// TIA Portal project "Pozycjoner_v7" (V15.1) (continued)
REGION Network 3: Line 1 is in or out range: 5mm around Y avg point
   #_w1 := #Enabled AND ((#Line1.Y1 < "DB_Average positions".Ranges.DiffX.Min) OR (#Line1.Y1 > "DB_Average positions".Ranges.DiffX.Max));
   IF #_w1 THEN #DiffResult := #Line1.Y1 - "DB_Average positions".AveragePosition.Y; END_IF;
   #SetCount1 := #_w1 AND NOT #Ptrig1;   // rising edge
   #Ptrig1 := #_w1;
   IF #Enabled AND ("DB_Average positions".Ranges.DiffX.Min <= #Line1.Y1) AND (#Line1.Y1 <= "DB_Average positions".Ranges.DiffX.Max) THEN
       #GeneralXavg := "DB_Drivers".X_AVG;
       #MoveToCenter_IR := TRUE;
   END_IF;
   IF #SetCount1 THEN
       #MainCounter := 1;
       #RECountLine3 := 0;
   END_IF;
END_REGION

REGION Network 4: Shift by difference value
   RUNG wire#powerrail
      { S7_Templates := "SrcType := Real" } GT_Contact(in1 := #DiffResult, in2 := 0.0)
      Sub(in1 := "DB_Average positions".AveragePosition.Y, in2 := #DiffResult, out => #ShiftDifValue)
   END_RUNG
   RUNG wire#powerrail
      { S7_Templates := "SrcType := Real" } LT_Contact(in1 := #DiffResult, in2 := 0.0)
      { S7_Templates := "SrcType := Real" } Abs(in := #DiffResult, out => #DiffResult)
      Add(in1 := "DB_Average positions".AveragePosition.Y, in2 := #DiffResult, out => #ShiftDifValue)
   END_RUNG
   // the same network as SCL:
   IF #DiffResult > 0.0 THEN
       #ShiftDifValue := "DB_Average positions".AveragePosition.Y - #DiffResult;
   END_IF;
   #_w1 := #DiffResult < 0.0;
   IF #_w1 THEN
       #DiffResult := ABS(#DiffResult);
       #ShiftDifValue := "DB_Average positions".AveragePosition.Y + #DiffResult;
   END_IF;
END_REGION

REGION Network 5: Movement to the new line: 3
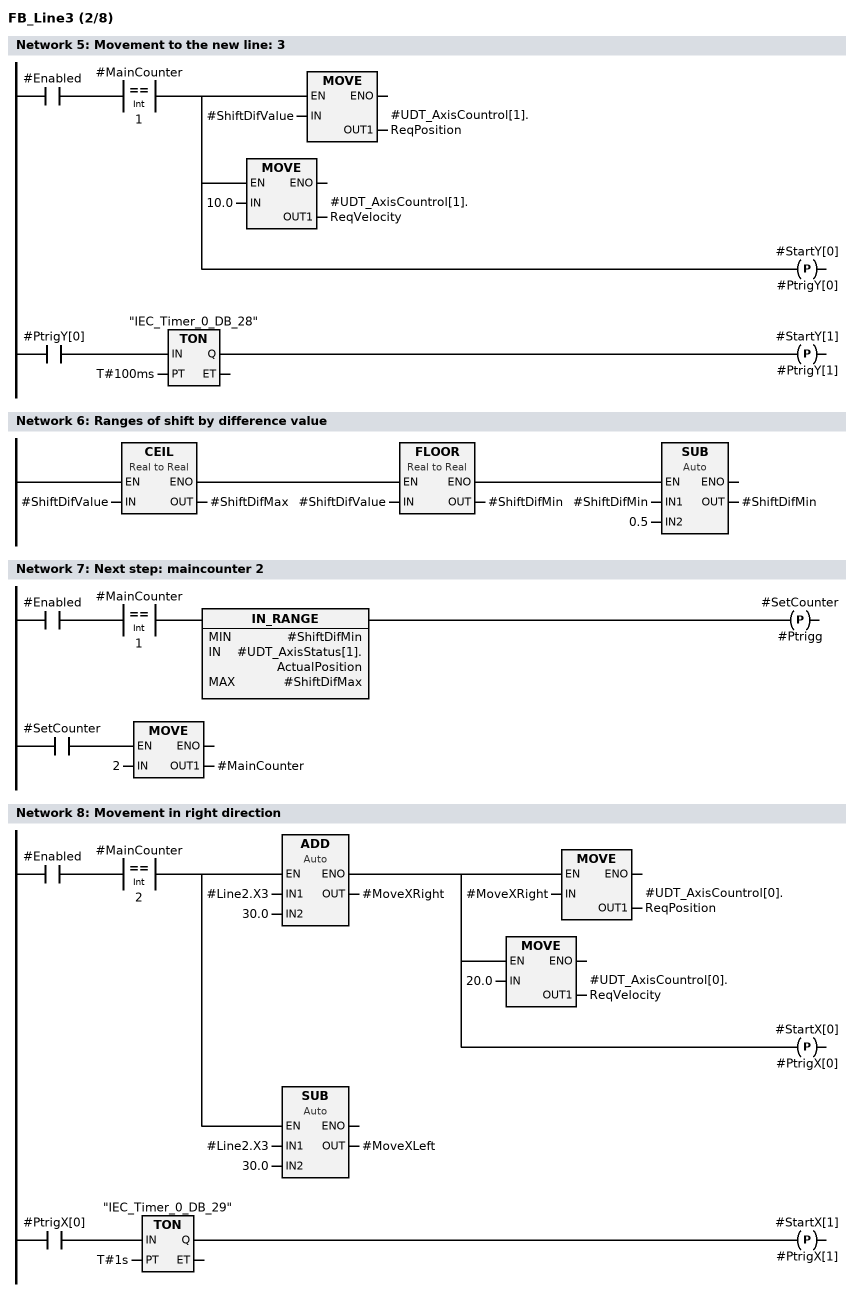
   #_w1 := #Enabled AND (#MainCounter = 1);
   IF #_w1 THEN
       #UDT_AxisCountrol[1].ReqPosition := #ShiftDifValue;
       #UDT_AxisCountrol[1].ReqVelocity := 10.0;
   END_IF;
   #StartY[0] := #_w1 AND NOT #PtrigY[0];   // rising edge
   #PtrigY[0] := #_w1;
   "IEC_Timer_0_DB_28".TON(IN := #PtrigY[0], PT := T#100ms);
   #StartY[1] := "IEC_Timer_0_DB_28".Q AND NOT #PtrigY[1];   // rising edge
   #PtrigY[1] := "IEC_Timer_0_DB_28".Q;
END_REGION

REGION Network 6: Ranges of shift by difference value
   #ShiftDifMax := CEIL(#ShiftDifValue);
   #ShiftDifMin := FLOOR(#ShiftDifValue);
   #ShiftDifMin := #ShiftDifMin - 0.5;
END_REGION

REGION Network 7: Next step: maincounter 2
   #_w1 := #Enabled AND (#MainCounter = 1) AND (#ShiftDifMin <= #UDT_AxisStatus[1].ActualPosition) AND (#UDT_AxisStatus[1].ActualPosition <= #ShiftDifMax);
   #SetCounter := #_w1 AND NOT #Ptrigg;   // rising edge
   #Ptrigg := #_w1;
   IF #SetCounter THEN #MainCounter := 2; END_IF;
END_REGION

REGION Network 8: Movement in right direction
   #_w1 := #Enabled AND (#MainCounter = 2);
   IF #_w1 THEN
       #MoveXRight := #Line2.X3 + 30.0;
       #UDT_AxisCountrol[0].ReqPosition := #MoveXRight;
       #UDT_AxisCountrol[0].ReqVelocity := 20.0;
   END_IF;
   #StartX[0] := #_w1 AND NOT #PtrigX[0];   // rising edge
   #PtrigX[0] := #_w1;
   IF #_w1 THEN #MoveXLeft := #Line2.X3 - 30.0; END_IF;
   "IEC_Timer_0_DB_29".TON(IN := #PtrigX[0], PT := T#1s);
   #StartX[1] := "IEC_Timer_0_DB_29".Q AND NOT #PtrigX[1];   // rising edge
   #PtrigX[1] := "IEC_Timer_0_DB_29".Q;
END_REGION

REGION Network 9: Stop movement
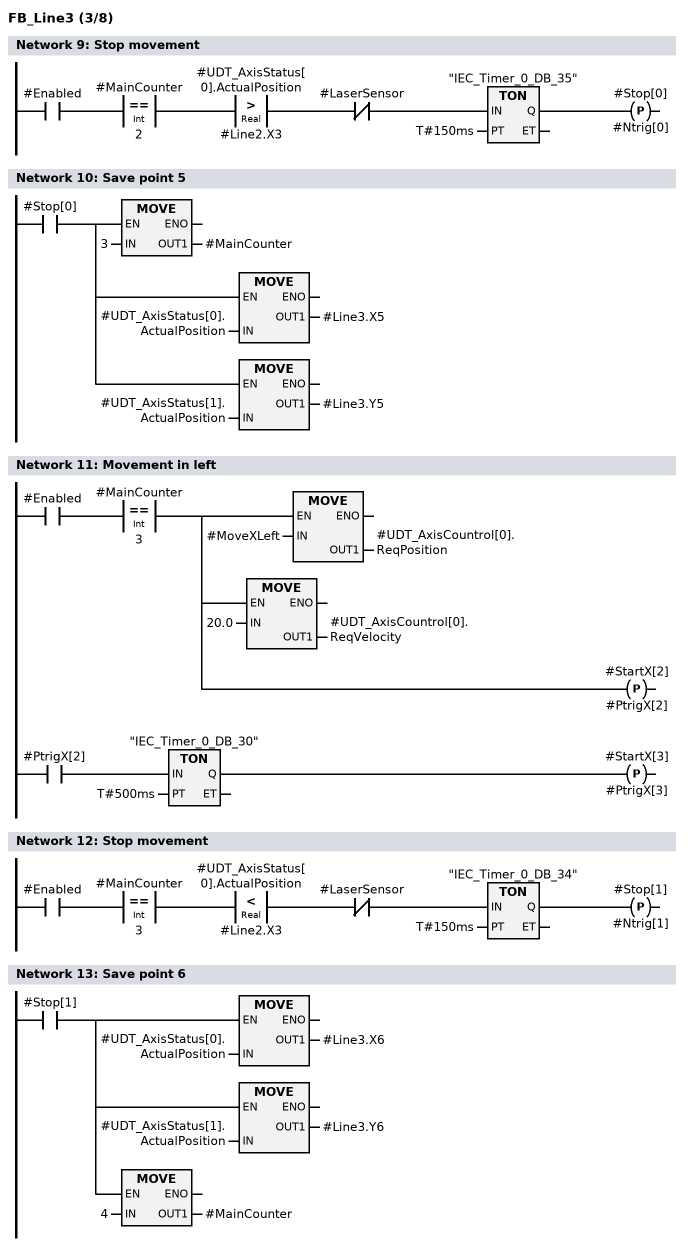
   "IEC_Timer_0_DB_35".TON(IN := #Enabled AND (#MainCounter = 2) AND (#UDT_AxisStatus[0].ActualPosition > #Line2.X3) AND NOT #LaserSensor,
                           PT := T#150ms);
   #Stop[0] := "IEC_Timer_0_DB_35".Q AND NOT #Ntrig[0];   // rising edge
   #Ntrig[0] := "IEC_Timer_0_DB_35".Q;
END_REGION

REGION Network 10: Save point 5
   RUNG wire#powerrail
      Contact( #Stop[0] )
      wire#w1
      Move(in := 3, out1 => #MainCounter)
   END_RUNG
   RUNG wire#w1
      Move(in := #UDT_AxisStatus[0].ActualPosition, out1 => #Line3.X5)
   END_RUNG
   RUNG wire#w1
      Move(in := #UDT_AxisStatus[1].ActualPosition, out1 => #Line3.Y5)
   END_RUNG
   // the same network as SCL:
   IF #Stop[0] THEN
       #MainCounter := 3;
       #Line3.X5 := #UDT_AxisStatus[0].ActualPosition;
       #Line3.Y5 := #UDT_AxisStatus[1].ActualPosition;
   END_IF;
END_REGION

REGION Network 11: Movement in left
   #_w1 := #Enabled AND (#MainCounter = 3);
   IF #_w1 THEN
       #UDT_AxisCountrol[0].ReqPosition := #MoveXLeft;
       #UDT_AxisCountrol[0].ReqVelocity := 20.0;
   END_IF;
   #StartX[2] := #_w1 AND NOT #PtrigX[2];   // rising edge
   #PtrigX[2] := #_w1;
   "IEC_Timer_0_DB_30".TON(IN := #PtrigX[2], PT := T#500ms);
   #StartX[3] := "IEC_Timer_0_DB_30".Q AND NOT #PtrigX[3];   // rising edge
   #PtrigX[3] := "IEC_Timer_0_DB_30".Q;
END_REGION

REGION Network 12: Stop movement
   "IEC_Timer_0_DB_34".TON(IN := #Enabled AND (#MainCounter = 3) AND (#UDT_AxisStatus[0].ActualPosition < #Line2.X3) AND NOT #LaserSensor,
                           PT := T#150ms);
   #Stop[1] := "IEC_Timer_0_DB_34".Q AND NOT #Ntrig[1];   // rising edge
   #Ntrig[1] := "IEC_Timer_0_DB_34".Q;
END_REGION

REGION Network 13: Save point 6
   RUNG wire#powerrail
      Contact( #Stop[1] )
      wire#w1
      Move(in := #UDT_AxisStatus[0].ActualPosition, out1 => #Line3.X6)
   END_RUNG
   RUNG wire#w1
      Move(in := #UDT_AxisStatus[1].ActualPosition, out1 => #Line3.Y6)
   END_RUNG
   RUNG wire#w1
      Move(in := 4, out1 => #MainCounter)
   END_RUNG
   // the same network as SCL:
   IF #Stop[1] THEN
       #Line3.X6 := #UDT_AxisStatus[0].ActualPosition;
       #Line3.Y6 := #UDT_AxisStatus[1].ActualPosition;
       #MainCounter := 4;
   END_IF;
END_REGION

REGION Network 14: Movement to the center point
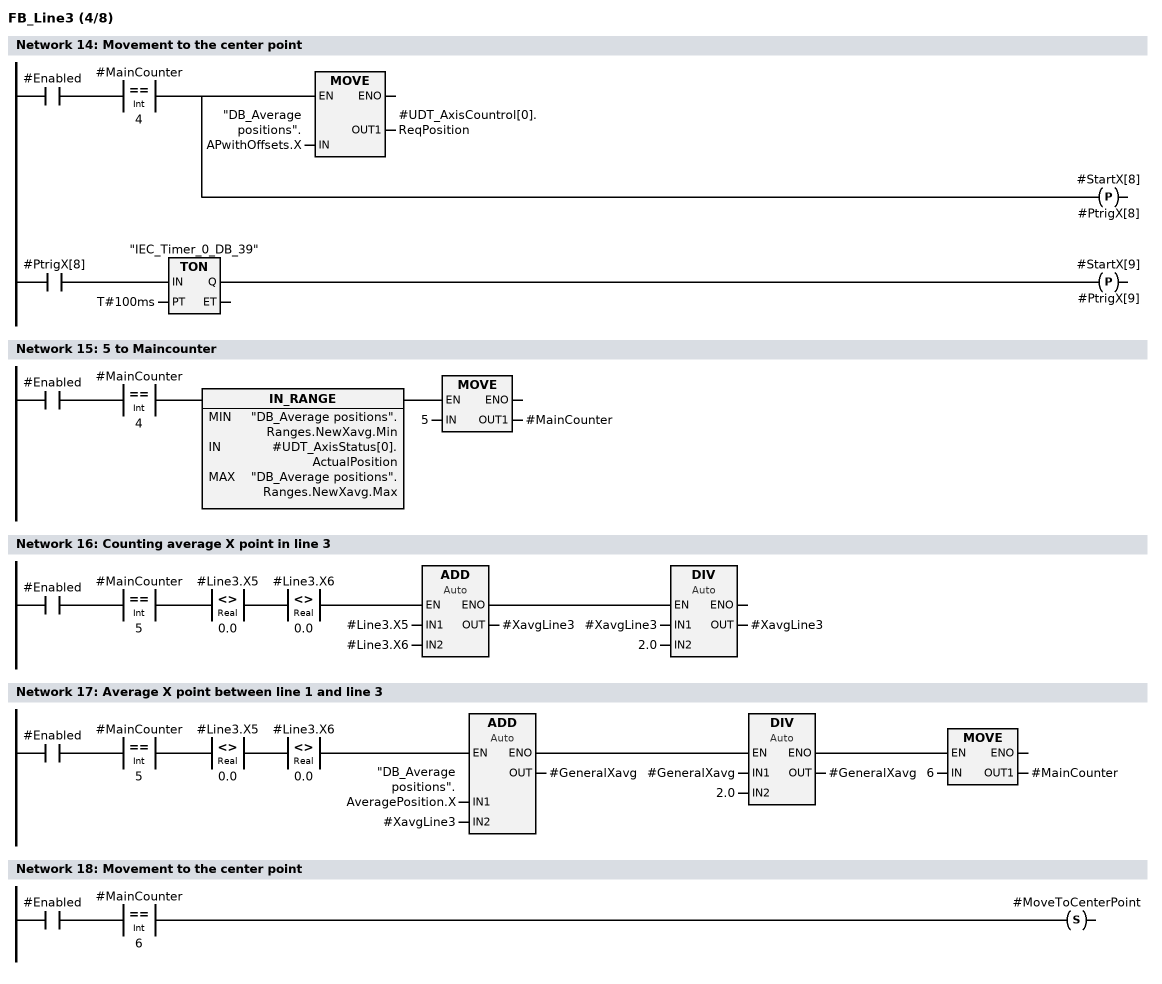
   #_w1 := #Enabled AND (#MainCounter = 4);
   IF #_w1 THEN #UDT_AxisCountrol[0].ReqPosition := "DB_Average positions".APwithOffsets.X; END_IF;
   #StartX[8] := #_w1 AND NOT #PtrigX[8];   // rising edge
   #PtrigX[8] := #_w1;
   "IEC_Timer_0_DB_39".TON(IN := #PtrigX[8], PT := T#100ms);
   #StartX[9] := "IEC_Timer_0_DB_39".Q AND NOT #PtrigX[9];   // rising edge
   #PtrigX[9] := "IEC_Timer_0_DB_39".Q;
END_REGION

REGION Network 15: 5 to Maincounter
   RUNG wire#powerrail
      Contact( #Enabled )
      { S7_Templates := "SrcType := Int" } EQ_Contact(in1 := #MainCounter, in2 := 4)
      { S7_Templates := "SrcType := Real" } InRange(min := "DB_Average positions".Ranges.NewXavg.Min, in := #UDT_AxisStatus[0].ActualPosition, max := "DB_Average positions".Ranges.NewXavg.Max)
      Move(in := 5, out1 => #MainCounter)
   END_RUNG
   // the same network as SCL:
   IF #Enabled AND (#MainCounter = 4) AND ("DB_Average positions".Ranges.NewXavg.Min <= #UDT_AxisStatus[0].ActualPosition) AND (#UDT_AxisStatus[0].ActualPosition <= "DB_Average positions".Ranges.NewXavg.Max) THEN
       #MainCounter := 5;
   END_IF;
END_REGION

REGION Network 16: Counting average X point in line 3
   RUNG wire#powerrail
      Contact( #Enabled )
      { S7_Templates := "SrcType := Int" } EQ_Contact(in1 := #MainCounter, in2 := 5)
      { S7_Templates := "SrcType := Real" } NE_Contact(in1 := #Line3.X5, in2 := 0.0)
      { S7_Templates := "SrcType := Real" } NE_Contact(in1 := #Line3.X6, in2 := 0.0)
      Add(in1 := #Line3.X5, in2 := #Line3.X6, out => #XavgLine3)
      Div(in1 := #XavgLine3, in2 := 2.0, out => #XavgLine3)
   END_RUNG
   // the same network as SCL:
   IF #Enabled AND (#MainCounter = 5) AND (#Line3.X5 <> 0.0) AND (#Line3.X6 <> 0.0) THEN
       #XavgLine3 := #Line3.X5 + #Line3.X6;
       #XavgLine3 := #XavgLine3 / 2.0;
   END_IF;
END_REGION

REGION Network 17: Average X point between line 1 and line 3
   RUNG wire#powerrail
      Contact( #Enabled )
      { S7_Templates := "SrcType := Int" } EQ_Contact(in1 := #MainCounter, in2 := 5)
      { S7_Templates := "SrcType := Real" } NE_Contact(in1 := #Line3.X5, in2 := 0.0)
      { S7_Templates := "SrcType := Real" } NE_Contact(in1 := #Line3.X6, in2 := 0.0)
      Add(in1 := "DB_Average positions".AveragePosition.X, in2 := #XavgLine3, out => #GeneralXavg)
      Div(in1 := #GeneralXavg, in2 := 2.0, out => #GeneralXavg)
      Move(in := 6, out1 => #MainCounter)
   END_RUNG
   // the same network as SCL:
   IF #Enabled AND (#MainCounter = 5) AND (#Line3.X5 <> 0.0) AND (#Line3.X6 <> 0.0) THEN
       #GeneralXavg := "DB_Average positions".AveragePosition.X + #XavgLine3;
       #GeneralXavg := #GeneralXavg / 2.0;
       #MainCounter := 6;
   END_IF;
END_REGION

REGION Network 18: Movement to the center point
   RUNG wire#powerrail
      Contact( #Enabled )
      { S7_Templates := "SrcType := Int" } EQ_Contact(in1 := #MainCounter, in2 := 6)
      S_Coil( #MoveToCenterPoint )
   END_RUNG
   // the same network as SCL:
   IF #Enabled AND (#MainCounter = 6) THEN #MoveToCenterPoint := TRUE; END_IF;
END_REGION

REGION Network 19: Movement to the center point
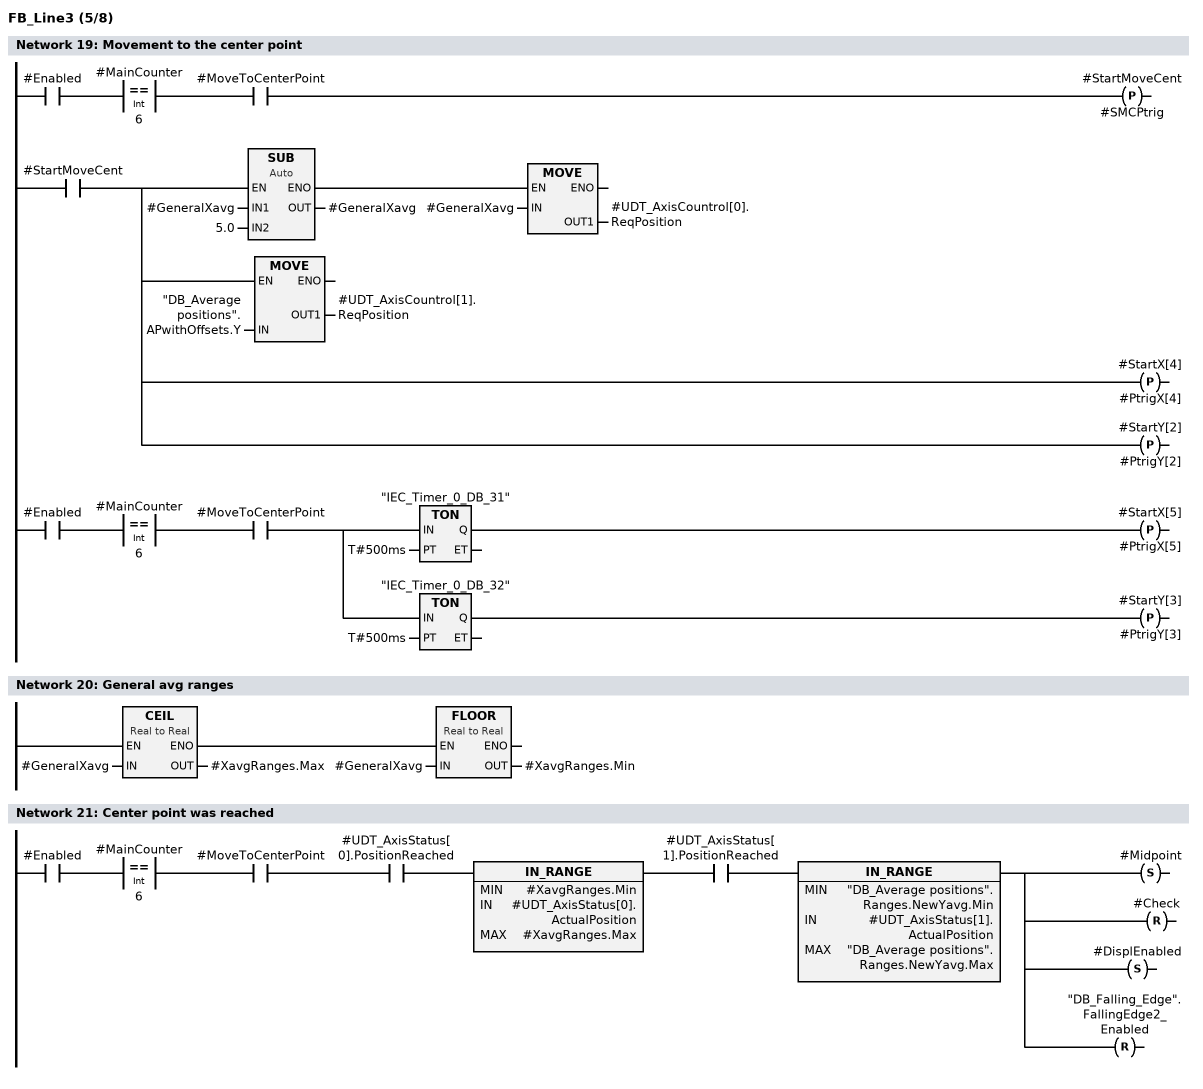
   #_w1 := #Enabled AND (#MainCounter = 6) AND #MoveToCenterPoint;
   #StartMoveCent := #_w1 AND NOT #SMCPtrig;   // rising edge
   #SMCPtrig := #_w1;
   IF #StartMoveCent THEN
       #GeneralXavg := #GeneralXavg - 5.0;
       #UDT_AxisCountrol[0].ReqPosition := #GeneralXavg;
       #UDT_AxisCountrol[1].ReqPosition := "DB_Average positions".APwithOffsets.Y;
   END_IF;
   #StartX[4] := #StartMoveCent AND NOT #PtrigX[4];   // rising edge
   #PtrigX[4] := #StartMoveCent;
   #StartY[2] := #StartMoveCent AND NOT #PtrigY[2];   // rising edge
   #PtrigY[2] := #StartMoveCent;
   #_w2 := #Enabled AND (#MainCounter = 6) AND #MoveToCenterPoint;
   "IEC_Timer_0_DB_31".TON(IN := #_w2, PT := T#500ms);
   #StartX[5] := "IEC_Timer_0_DB_31".Q AND NOT #PtrigX[5];   // rising edge
   #PtrigX[5] := "IEC_Timer_0_DB_31".Q;
   "IEC_Timer_0_DB_32".TON(IN := #_w2, PT := T#500ms);
   #StartY[3] := "IEC_Timer_0_DB_32".Q AND NOT #PtrigY[3];   // rising edge
   #PtrigY[3] := "IEC_Timer_0_DB_32".Q;
END_REGION

REGION Network 20: General avg ranges
   #XavgRanges.Max := CEIL(#GeneralXavg);
   #XavgRanges.Min := FLOOR(#GeneralXavg);
END_REGION

REGION Network 21: Center point was reached
   RUNG wire#powerrail
      Contact( #Enabled )
      { S7_Templates := "SrcType := Int" } EQ_Contact(in1 := #MainCounter, in2 := 6)
      Contact( #MoveToCenterPoint )
      Contact( #UDT_AxisStatus[0].PositionReached )
      { S7_Templates := "SrcType := Real" } InRange(min := #XavgRanges.Min, in := #UDT_AxisStatus[0].ActualPosition, max := #XavgRanges.Max)
      Contact( #UDT_AxisStatus[1].PositionReached )
      { S7_Templates := "SrcType := Real" } InRange(min := "DB_Average positions".Ranges.NewYavg.Min, in := #UDT_AxisStatus[1].ActualPosition, max := "DB_Average positions".Ranges.NewYavg.Max)
      wire#w1
      S_Coil( #Midpoint )
   END_RUNG
   RUNG wire#w1
      R_Coil( #Check )
   END_RUNG
   RUNG wire#w1
      S_Coil( #DisplEnabled )
   END_RUNG
   RUNG wire#w1
      R_Coil( "DB_Falling_Edge".FallingEdge2_Enabled )
   END_RUNG
   // the same network as SCL:
   IF #Enabled AND (#MainCounter = 6) AND #MoveToCenterPoint AND #UDT_AxisStatus[0].PositionReached AND (#XavgRanges.Min <= #UDT_AxisStatus[0].ActualPosition) AND (#UDT_AxisStatus[0].ActualPosition <= #XavgRanges.Max) AND #UDT_AxisStatus[1].PositionReached AND ("DB_Average positions".Ranges.NewYavg.Min <= #UDT_AxisStatus[1].ActualPosition) AND (#UDT_AxisStatus[1].ActualPosition <= "DB_Average positions".Ranges.NewYavg.Max) THEN
       #Midpoint := TRUE;
       #Check := FALSE;
       #DisplEnabled := TRUE;
       "DB_Falling_Edge".FallingEdge2_Enabled := FALSE;
   END_IF;
END_REGION

REGION Network 22: Line 1 is IN 5mm range, movement to the center point without making line 3
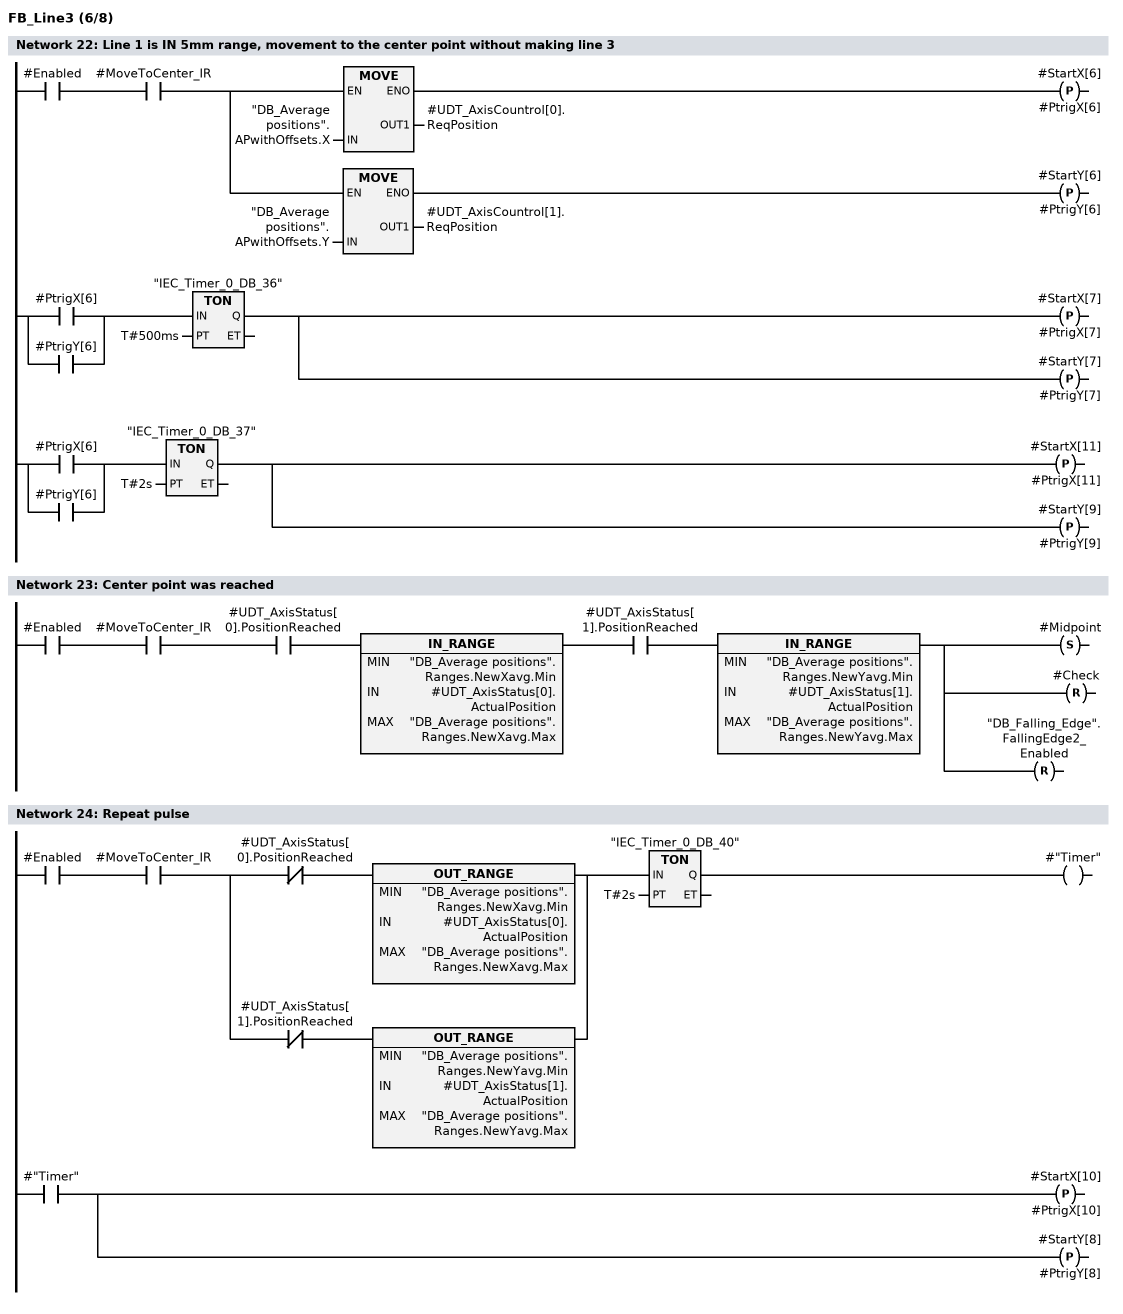
   #_w1 := #Enabled AND #MoveToCenter_IR;
   IF #_w1 THEN #UDT_AxisCountrol[0].ReqPosition := "DB_Average positions".APwithOffsets.X; END_IF;
   #StartX[6] := #_w1 AND NOT #PtrigX[6];   // rising edge
   #PtrigX[6] := #_w1;
   IF #_w1 THEN #UDT_AxisCountrol[1].ReqPosition := "DB_Average positions".APwithOffsets.Y; END_IF;
   #StartY[6] := #_w1 AND NOT #PtrigY[6];   // rising edge
   #PtrigY[6] := #_w1;
   "IEC_Timer_0_DB_36".TON(IN := #PtrigX[6] OR #PtrigY[6], PT := T#500ms);
   #StartX[7] := "IEC_Timer_0_DB_36".Q AND NOT #PtrigX[7];   // rising edge
   #PtrigX[7] := "IEC_Timer_0_DB_36".Q;
   #StartY[7] := "IEC_Timer_0_DB_36".Q AND NOT #PtrigY[7];   // rising edge
   #PtrigY[7] := "IEC_Timer_0_DB_36".Q;
   "IEC_Timer_0_DB_37".TON(IN := #PtrigX[6] OR #PtrigY[6], PT := T#2s);
   #StartX[11] := "IEC_Timer_0_DB_37".Q AND NOT #PtrigX[11];   // rising edge
   #PtrigX[11] := "IEC_Timer_0_DB_37".Q;
   #StartY[9] := "IEC_Timer_0_DB_37".Q AND NOT #PtrigY[9];   // rising edge
   #PtrigY[9] := "IEC_Timer_0_DB_37".Q;
END_REGION

REGION Network 23: Center point was reached
   RUNG wire#powerrail
      Contact( #Enabled )
      Contact( #MoveToCenter_IR )
      Contact( #UDT_AxisStatus[0].PositionReached )
      { S7_Templates := "SrcType := Real" } InRange(min := "DB_Average positions".Ranges.NewXavg.Min, in := #UDT_AxisStatus[0].ActualPosition, max := "DB_Average positions".Ranges.NewXavg.Max)
      Contact( #UDT_AxisStatus[1].PositionReached )
      { S7_Templates := "SrcType := Real" } InRange(min := "DB_Average positions".Ranges.NewYavg.Min, in := #UDT_AxisStatus[1].ActualPosition, max := "DB_Average positions".Ranges.NewYavg.Max)
      wire#w1
      S_Coil( #Midpoint )
   END_RUNG
   RUNG wire#w1
      R_Coil( #Check )
   END_RUNG
   RUNG wire#w1
      R_Coil( "DB_Falling_Edge".FallingEdge2_Enabled )
   END_RUNG
   // the same network as SCL:
   IF #Enabled AND #MoveToCenter_IR AND #UDT_AxisStatus[0].PositionReached AND ("DB_Average positions".Ranges.NewXavg.Min <= #UDT_AxisStatus[0].ActualPosition) AND (#UDT_AxisStatus[0].ActualPosition <= "DB_Average positions".Ranges.NewXavg.Max) AND #UDT_AxisStatus[1].PositionReached AND ("DB_Average positions".Ranges.NewYavg.Min <= #UDT_AxisStatus[1].ActualPosition) AND (#UDT_AxisStatus[1].ActualPosition <= "DB_Average positions".Ranges.NewYavg.Max) THEN
       #Midpoint := TRUE;
       #Check := FALSE;
       "DB_Falling_Edge".FallingEdge2_Enabled := FALSE;
   END_IF;
END_REGION

REGION Network 24: Repeat pulse
   "IEC_Timer_0_DB_40".TON(IN := #Enabled AND #MoveToCenter_IR AND ((NOT #UDT_AxisStatus[0].PositionReached AND ((#UDT_AxisStatus[0].ActualPosition < "DB_Average positions".Ranges.NewXavg.Min) OR (#UDT_AxisStatus[0].ActualPosition > "DB_Average positions".Ranges.NewXavg.Max))) OR (NOT #UDT_AxisStatus[1].PositionReached AND ((#UDT_AxisStatus[1].ActualPosition < "DB_Average positions".Ranges.NewYavg.Min) OR (#UDT_AxisStatus[1].ActualPosition > "DB_Average positions".Ranges.NewYavg.Max)))),
                           PT := T#2s);
   #"Timer" := "IEC_Timer_0_DB_40".Q;
   #StartX[10] := #"Timer" AND NOT #PtrigX[10];   // rising edge
   #PtrigX[10] := #"Timer";
   #StartY[8] := #"Timer" AND NOT #PtrigY[8];   // rising edge
   #PtrigY[8] := #"Timer";
END_REGION

REGION Network 25: Start Movement Command
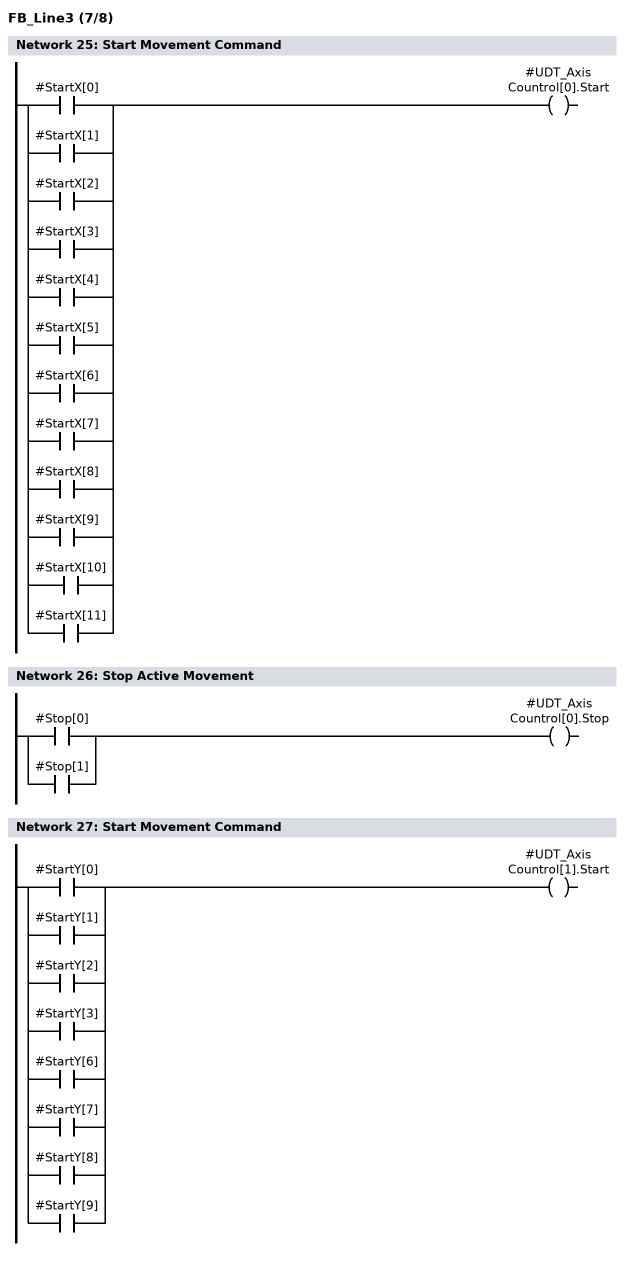
   RUNG wire#powerrail
      Contact( #StartX[0] )
      wire#w1
      Coil( #UDT_AxisCountrol[0].Start )
   END_RUNG
   RUNG wire#powerrail
      Contact( #StartX[1] )
   END_RUNG wire#w1
   RUNG wire#powerrail
      Contact( #StartX[2] )
   END_RUNG wire#w1
   RUNG wire#powerrail
      Contact( #StartX[3] )
   END_RUNG wire#w1
   RUNG wire#powerrail
      Contact( #StartX[4] )
   END_RUNG wire#w1
   RUNG wire#powerrail
      Contact( #StartX[5] )
   END_RUNG wire#w1
   RUNG wire#powerrail
      Contact( #StartX[6] )
   END_RUNG wire#w1
   RUNG wire#powerrail
      Contact( #StartX[7] )
   END_RUNG wire#w1
   RUNG wire#powerrail
      Contact( #StartX[8] )
   END_RUNG wire#w1
   RUNG wire#powerrail
      Contact( #StartX[9] )
   END_RUNG wire#w1
   RUNG wire#powerrail
      Contact( #StartX[10] )
   END_RUNG wire#w1
   RUNG wire#powerrail
      Contact( #StartX[11] )
   END_RUNG wire#w1
   // the same network as SCL:
   #UDT_AxisCountrol[0].Start := #StartX[0] OR #StartX[1] OR #StartX[2] OR #StartX[3] OR #StartX[4] OR #StartX[5] OR #StartX[6] OR #StartX[7] OR #StartX[8] OR #StartX[9] OR #StartX[10] OR #StartX[11];
END_REGION

REGION Network 26: Stop Active Movement
   RUNG wire#powerrail
      Contact( #Stop[0] )
      wire#w1
      Coil( #UDT_AxisCountrol[0].Stop )
   END_RUNG
   RUNG wire#powerrail
      Contact( #Stop[1] )
   END_RUNG wire#w1
   // the same network as SCL:
   #UDT_AxisCountrol[0].Stop := #Stop[0] OR #Stop[1];
END_REGION

REGION Network 27: Start Movement Command
   RUNG wire#powerrail
      Contact( #StartY[0] )
      wire#w1
      Coil( #UDT_AxisCountrol[1].Start )
   END_RUNG
   RUNG wire#powerrail
      Contact( #StartY[1] )
   END_RUNG wire#w1
   RUNG wire#powerrail
      Contact( #StartY[2] )
   END_RUNG wire#w1
   RUNG wire#powerrail
      Contact( #StartY[3] )
   END_RUNG wire#w1
   RUNG wire#powerrail
      Contact( #StartY[6] )
   END_RUNG wire#w1
   RUNG wire#powerrail
      Contact( #StartY[7] )
   END_RUNG wire#w1
   RUNG wire#powerrail
      Contact( #StartY[8] )
   END_RUNG wire#w1
   RUNG wire#powerrail
      Contact( #StartY[9] )
   END_RUNG wire#w1
   // the same network as SCL:
   #UDT_AxisCountrol[1].Start := #StartY[0] OR #StartY[1] OR #StartY[2] OR #StartY[3] OR #StartY[6] OR #StartY[7] OR #StartY[8] OR #StartY[9];
END_REGION

REGION Network 28: Save points
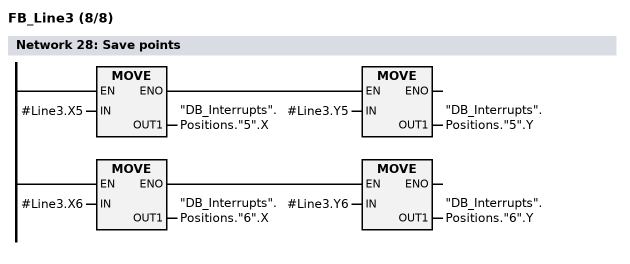
   RUNG wire#powerrail
      Move(in := #Line3.X5, out1 => "DB_Interrupts".Positions."5".X)
      Move(in := #Line3.Y5, out1 => "DB_Interrupts".Positions."5".Y)
   END_RUNG
   RUNG wire#powerrail
      Move(in := #Line3.X6, out1 => "DB_Interrupts".Positions."6".X)
      Move(in := #Line3.Y6, out1 => "DB_Interrupts".Positions."6".Y)
   END_RUNG
   // the same network as SCL:
   "DB_Interrupts".Positions."5".X := #Line3.X5;
   "DB_Interrupts".Positions."5".Y := #Line3.Y5;
   "DB_Interrupts".Positions."6".X := #Line3.X6;
   "DB_Interrupts".Positions."6".Y := #Line3.Y6;
END_REGION
END_FUNCTION_BLOCK

// folder: Displacement/Object displacement

FUNCTION_BLOCK "FB_Displacement"   // FB15, LAD
{ S7_Optimized_Access := 'TRUE' }
VERSION : 0.1
   VAR
      UDT_AxisControl : Array[0..2] of "UDT_AxisControl";
      UDT_AxisStatus : Array[0..2] of "UDT_AxisStatus";
      MainCounter : Int;   // Main couner - indicate which part of program is active
      StartX : Array[0..3] of Bool;   // Start X pulse
      PTrigX : Array[0..3] of Bool;   // X ptrig - previous state
      StartY : Array[0..3] of Bool;   // Start Y pulse
      PTrigY : Array[0..3] of Bool;   // Y ptrig - previous state
      StartZ : Array[0..10] of Bool;   // Start Z pulse
      PtrigZ : Array[0..10] of Bool;   // Z ptrig - previous state
      Electromagnet : Bool;   // Electromagnet variable
      DiplacementMode : Bool;   // Enable/disable this mode as active
      Ptrig : Bool;   // Additional variable
      ZOffset : Real;   // Z offset between CW limit and item
      ZMedPos : Real;   // Z position, half of CCW limit
      Zmin : Int;   // Z min range: ZOffset
      Zmax : Int;   // Z max range: ZOffset
      ZminMP : Int;   // Z min range: ZMedPos
      ZmaxMP : Int;   // Z max range: ZMedPos
      ZOfsmax : Real;   // 2 mm above Z offset value
      TpY : Real;   // Target position in Y axis
      TpX : Real;   // Target position in X axis
      SensorPos : Struct   // Available sensor coordinates
         XPos : Real;
         YPos : Real;
         SensNumb : Int;
      END_STRUCT;
      SensorRanges : Struct   // Available sensor ranges
         Xmin : Real;
         Xmax : Real;
         Ymin : Real;
         Ymax : Real;
      END_STRUCT;
      Vx : Real;   // X velocity
      Vy : Real;   // Y velocity
      HalfS : Real;   // Half of the distance
      PlaceOcup : Struct   // Place ocuppied for each sensor
         Sens1 : Bool;
         Sens2 : Bool;
         Sens3 : Bool;
         Sens4 : Bool;
         Place : Int;
      END_STRUCT;
      X_out_min : Int;   // X min range of the previous position
      X_out_max : Int;   // X max range of the previous position
      Y_out_min : Int;
      Y_out_max : Int;
      TargetPosition : Bool;   // Target position (previous position - before interrupt was started)
      Tim : Array[0..8] of Bool;   // Additional timers
      StopEM : Bool;
      Ntrig : Bool;
      Sz : Real;   // Z distance
      Vz : Real;   // Z velocity
      TpRanges : Struct
         Min : Real;
         Max : Real;
      END_STRUCT;
   END_VAR
   VAR CONSTANT
      false : Bool;
   END_VAR
   VAR_TEMP   // added for the SCL form of the ladder/FBD networks
      _w1 : Bool;
   END_VAR
BEGIN

REGION Network 1: Enabled mode
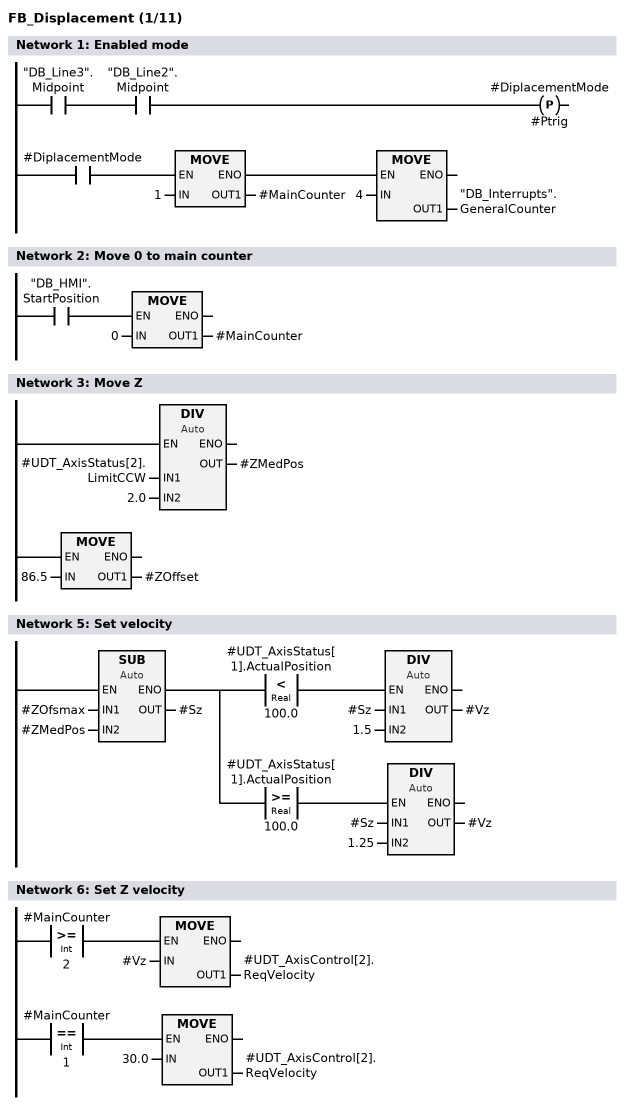
   #_w1 := "DB_Line3".Midpoint AND "DB_Line2".Midpoint;
   #DiplacementMode := #_w1 AND NOT #Ptrig;   // rising edge
   #Ptrig := #_w1;
   IF #DiplacementMode THEN
       #MainCounter := 1;
       "DB_Interrupts".GeneralCounter := 4;
   END_IF;
END_REGION

REGION Network 2: Move 0 to main counter
   RUNG wire#powerrail
      Contact( "DB_HMI".StartPosition )
      Move(in := 0, out1 => #MainCounter)
   END_RUNG
   // the same network as SCL:
   IF "DB_HMI".StartPosition THEN #MainCounter := 0; END_IF;
END_REGION

REGION Network 3: Move Z
   RUNG wire#powerrail
      Div(in1 := #UDT_AxisStatus[2].LimitCCW, in2 := 2.0, out => #ZMedPos)
   END_RUNG
   RUNG wire#powerrail
      Move(in := 86.5, out1 => #ZOffset)
   END_RUNG
   // the same network as SCL:
   #ZMedPos := #UDT_AxisStatus[2].LimitCCW / 2.0;
   #ZOffset := 86.5;
END_REGION

REGION Network 5: Set velocity
   RUNG wire#powerrail
      Sub(in1 := #ZOfsmax, in2 := #ZMedPos, out => #Sz)
      wire#w1
      { S7_Templates := "SrcType := Real" } LT_Contact(in1 := #UDT_AxisStatus[1].ActualPosition, in2 := 100.0)
      Div(in1 := #Sz, in2 := 1.5, out => #Vz)
   END_RUNG
   RUNG wire#w1
      { S7_Templates := "SrcType := Real" } GE_Contact(in1 := #UDT_AxisStatus[1].ActualPosition, in2 := 100.0)
      Div(in1 := #Sz, in2 := 1.25, out => #Vz)
   END_RUNG
   // the same network as SCL:
   #Sz := #ZOfsmax - #ZMedPos;
   IF #UDT_AxisStatus[1].ActualPosition < 100.0 THEN #Vz := #Sz / 1.5; END_IF;
   IF #UDT_AxisStatus[1].ActualPosition >= 100.0 THEN #Vz := #Sz / 1.25; END_IF;
END_REGION

REGION Network 6: Set Z velocity
   RUNG wire#powerrail
      { S7_Templates := "SrcType := Int" } GE_Contact(in1 := #MainCounter, in2 := 2)
      Move(in := #Vz, out1 => #UDT_AxisControl[2].ReqVelocity)
   END_RUNG
   RUNG wire#powerrail
      { S7_Templates := "SrcType := Int" } EQ_Contact(in1 := #MainCounter, in2 := 1)
      Move(in := 30.0, out1 => #UDT_AxisControl[2].ReqVelocity)
   END_RUNG
   // the same network as SCL:
   IF #MainCounter >= 2 THEN #UDT_AxisControl[2].ReqVelocity := #Vz; END_IF;
   IF #MainCounter = 1 THEN #UDT_AxisControl[2].ReqVelocity := 30.0; END_IF;
END_REGION

REGION Network 7: Grab item
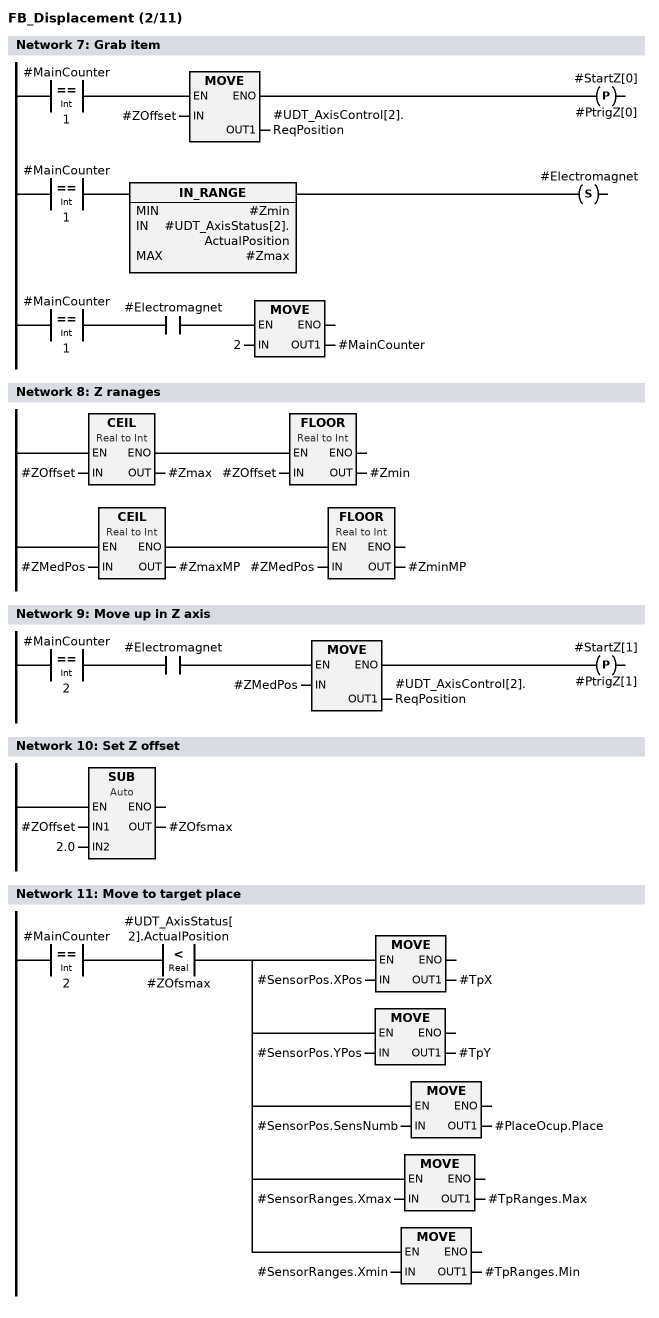
   #_w1 := #MainCounter = 1;
   IF #_w1 THEN #UDT_AxisControl[2].ReqPosition := #ZOffset; END_IF;
   #StartZ[0] := #_w1 AND NOT #PtrigZ[0];   // rising edge
   #PtrigZ[0] := #_w1;
   IF (#MainCounter = 1) AND (#Zmin <= #UDT_AxisStatus[2].ActualPosition) AND (#UDT_AxisStatus[2].ActualPosition <= #Zmax) THEN
       #Electromagnet := TRUE;
   END_IF;
   IF (#MainCounter = 1) AND #Electromagnet THEN #MainCounter := 2; END_IF;
END_REGION

REGION Network 8: Z ranages
   #Zmax := CEIL(#ZOffset);
   #Zmin := FLOOR(#ZOffset);
   #ZmaxMP := CEIL(#ZMedPos);
   #ZminMP := FLOOR(#ZMedPos);
END_REGION

REGION Network 9: Move up in Z axis
   #_w1 := (#MainCounter = 2) AND #Electromagnet;
   IF #_w1 THEN #UDT_AxisControl[2].ReqPosition := #ZMedPos; END_IF;
   #StartZ[1] := #_w1 AND NOT #PtrigZ[1];   // rising edge
   #PtrigZ[1] := #_w1;
END_REGION

REGION Network 10: Set Z offset
   RUNG wire#powerrail
      Sub(in1 := #ZOffset, in2 := 2.0, out => #ZOfsmax)
   END_RUNG
   // the same network as SCL:
   #ZOfsmax := #ZOffset - 2.0;
END_REGION

REGION Network 11: Move to target place
   RUNG wire#powerrail
      { S7_Templates := "SrcType := Int" } EQ_Contact(in1 := #MainCounter, in2 := 2)
      { S7_Templates := "SrcType := Real" } LT_Contact(in1 := #UDT_AxisStatus[2].ActualPosition, in2 := #ZOfsmax)
      wire#w1
      Move(in := #SensorPos.XPos, out1 => #TpX)
   END_RUNG
   RUNG wire#w1
      Move(in := #SensorPos.YPos, out1 => #TpY)
   END_RUNG
   RUNG wire#w1
      Move(in := #SensorPos.SensNumb, out1 => #PlaceOcup.Place)
   END_RUNG
   RUNG wire#w1
      Move(in := #SensorRanges.Xmax, out1 => #TpRanges.Max)
   END_RUNG
   RUNG wire#w1
      Move(in := #SensorRanges.Xmin, out1 => #TpRanges.Min)
   END_RUNG
   // the same network as SCL:
   IF (#MainCounter = 2) AND (#UDT_AxisStatus[2].ActualPosition < #ZOfsmax) THEN
       #TpX := #SensorPos.XPos;
       #TpY := #SensorPos.YPos;
       #PlaceOcup.Place := #SensorPos.SensNumb;
       #TpRanges.Max := #SensorRanges.Xmax;
       #TpRanges.Min := #SensorRanges.Xmin;
   END_IF;
END_REGION

REGION Network 12: Count velocity
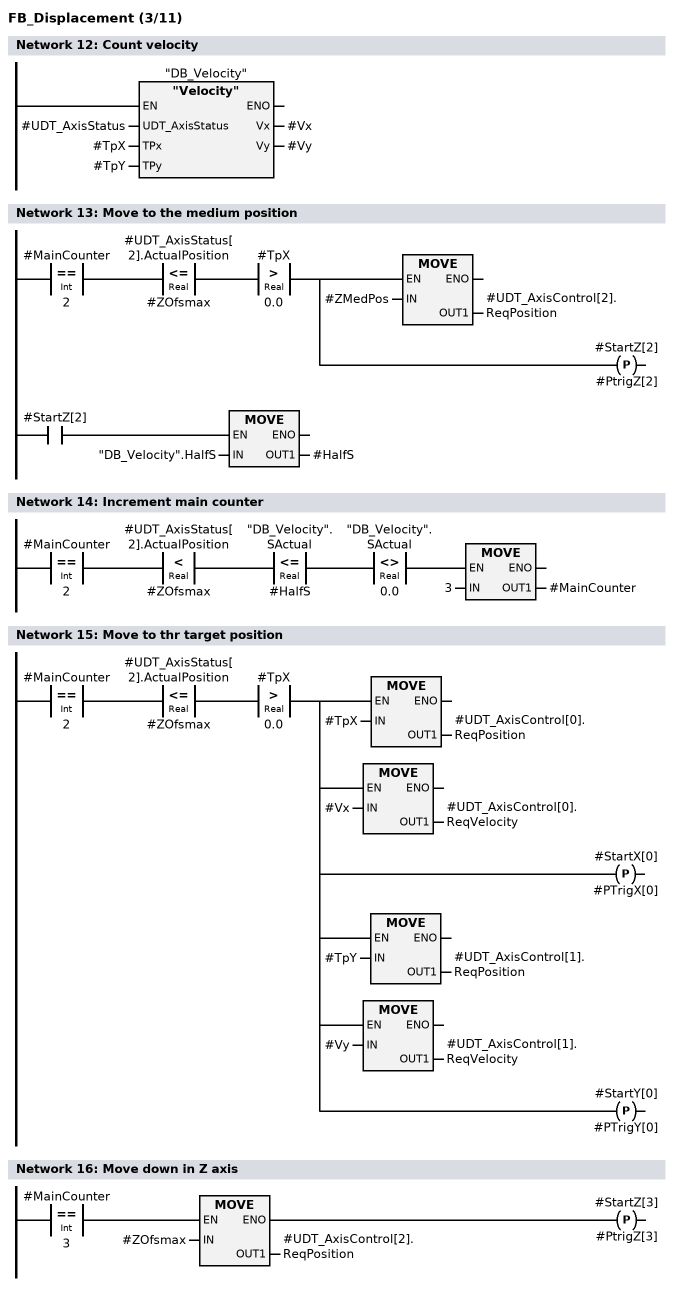
   RUNG wire#powerrail
      "DB_Velocity"(UDT_AxisStatus := #UDT_AxisStatus, TPx := #TpX, TPy := #TpY, Vx => #Vx, Vy => #Vy)
   END_RUNG
   // the same network as SCL:
   "DB_Velocity"(UDT_AxisStatus := #UDT_AxisStatus, TPx := #TpX, TPy := #TpY, Vx => #Vx, Vy => #Vy);   // "Velocity"
END_REGION

REGION Network 13: Move to the medium position
   #_w1 := (#MainCounter = 2) AND (#UDT_AxisStatus[2].ActualPosition <= #ZOfsmax) AND (#TpX > 0.0);
   IF #_w1 THEN #UDT_AxisControl[2].ReqPosition := #ZMedPos; END_IF;
   #StartZ[2] := #_w1 AND NOT #PtrigZ[2];   // rising edge
   #PtrigZ[2] := #_w1;
   IF #StartZ[2] THEN #HalfS := "DB_Velocity".HalfS; END_IF;
END_REGION

REGION Network 14: Increment main counter
   RUNG wire#powerrail
      { S7_Templates := "SrcType := Int" } EQ_Contact(in1 := #MainCounter, in2 := 2)
      { S7_Templates := "SrcType := Real" } LT_Contact(in1 := #UDT_AxisStatus[2].ActualPosition, in2 := #ZOfsmax)
      { S7_Templates := "SrcType := Real" } LE_Contact(in1 := "DB_Velocity".SActual, in2 := #HalfS)
      { S7_Templates := "SrcType := Real" } NE_Contact(in1 := "DB_Velocity".SActual, in2 := 0.0)
      Move(in := 3, out1 => #MainCounter)
   END_RUNG
   // the same network as SCL:
   IF (#MainCounter = 2) AND (#UDT_AxisStatus[2].ActualPosition < #ZOfsmax) AND ("DB_Velocity".SActual <= #HalfS) AND ("DB_Velocity".SActual <> 0.0) THEN
       #MainCounter := 3;
   END_IF;
END_REGION

REGION Network 15: Move to thr target position
   #_w1 := (#MainCounter = 2) AND (#UDT_AxisStatus[2].ActualPosition <= #ZOfsmax) AND (#TpX > 0.0);
   IF #_w1 THEN
       #UDT_AxisControl[0].ReqPosition := #TpX;
       #UDT_AxisControl[0].ReqVelocity := #Vx;
   END_IF;
   #StartX[0] := #_w1 AND NOT #PTrigX[0];   // rising edge
   #PTrigX[0] := #_w1;
   IF #_w1 THEN
       #UDT_AxisControl[1].ReqPosition := #TpY;
       #UDT_AxisControl[1].ReqVelocity := #Vy;
   END_IF;
   #StartY[0] := #_w1 AND NOT #PTrigY[0];   // rising edge
   #PTrigY[0] := #_w1;
END_REGION

REGION Network 16: Move down in Z axis
   #_w1 := #MainCounter = 3;
   IF #_w1 THEN #UDT_AxisControl[2].ReqPosition := #ZOfsmax; END_IF;
   #StartZ[3] := #_w1 AND NOT #PtrigZ[3];   // rising edge
   #PtrigZ[3] := #_w1;
END_REGION

REGION Network 17: Put the item
